screen "Balast Water Treatment Plant" 1280x800, template "Template"
   on GenerateScreen: "User_Change"(); "TitleUpdater"()
   Button "HmiScreenItemData_1" at 1,1 size 150x40; TextOn 'Back'; TextOff 'Main Index'
      on Release: ActivateScreen("02 Main Index", 0)
   TextField "Text field_63" at 383,107 size 72x30; Text 'Pre Dwell Time'
   Circle "Circle_29" at 1047,85 size 20x20
      Appearance <- "2102_TIME_CALCS_DB_POST_DWELL_TMR_DN"
   Button "HmiScreenItemData_9" at 10,60 size 158x27; TextOn 'Back'; TextOff 'BWTS Control'
   Button "HmiScreenItemData_4" at 14,150 size 75x47; TextOn 'Back'; TextOff 'Stop'; Authorization "Operate"
      on Release: function_efd93a16("BWTS Stop Confirm", 300, 200, -1, -1, 1)
      ObjectEnable <- "82_To_HMI_CRNT_MODE_GCU"
   Circle "Circle_20" at 137,105 size 29x29
      Appearance <- "80_From_HMI_RUN_IGG(1)"
   Button "HmiScreenItemData_3" at 14,93 size 75x47; TextOn 'Back'; TextOff 'Start'; Authorization "Operate"
      on Release: function_efd93a16("BWTS Start Confirm", 300, 200, -1, -1, 1)
      ObjectEnable <- "82_To_HMI_CRNT_MODE_GCU"
   Button "HmiScreenItemData_2" at 1129,1 size 150x40; TextOn 'Back'; TextOff 'BWTS Setup'
      on Release: ActivateScreen("Balast Water Treatment Setup", 0)
   TextField "Text field_1" at 290,107 size 68x30; Text 'Tank Selected'
   TextField "Text field_2" at 841,107 size 61x30; Text 'BWTS Started'
   TextField "Text field_3" at 568,107 size 62x30; Text 'IGGS Started'
   TextField "Text field_4" at 659,107 size 60x30; Text 'GCU Started'
   TextField "Text field_5" at 748,107 size 61x30; Text 'PGC Started'
   TextField "Text field_6" at 908,107 size 102x30; Text 'Gas Transfer Started'
   Circle "Circle_10" at 956,89 size 14x14
      Appearance <- "2110_BTCS_CNTRL_DB_BTCS_STEP"
   TextField "Text field_7" at 995,107 size 125x30; Text 'Treatment Cycle Completed'
   TextField "Text field_21" at 306,401 size 54x20; Text 'Closed'
      Visibility <- "20_TANKS_IP_DATA_RIO_06_FIRST_TANK_GTT_ISOL_VALVE_CLSD"
   TextField "Text field_22" at 306,401 size 54x20; Text 'Opened'
      Visibility <- "20_TANKS_IP_DATA_RIO_06_FIRST_TANK_GTT_ISOL_VALVE_OPEN"
   GraphicView "Graphic view_10" at 283,396 size 22x31; Picture "Graphic_162"
   TextField "Text field_25" at 306,482 size 54x20; Text 'Closed'
      Visibility <- "20_TANKS_IP_DATA_RIO_06_SECOND_TANK_GTT_ISOL_VALVE_CLSD"
   TextField "Text field_26" at 306,482 size 54x20; Text 'Opened'
      Visibility <- "20_TANKS_IP_DATA_RIO_06_SECOND_TANK_GTT_ISOL_VALVE_OPEN"
   IOField "I/O field_2" at 309,560 size 72x20; FormatPattern 999; Unit Nm³/hr
      ProcessValue <- "20_TANKS_IP_DATA_RIO_06_SECOND_TANK_USD_FLOW"
   IOField "I/O field_4" at 309,599 size 72x20; FormatPattern 999; Unit Nm³/hr
      ProcessValue <- "20_TANKS_IP_DATA_RIO_06_SECOND_TANK_MBG_FLOW"
   TextField "Text field_27" at 263,602 size 29x14; Text 'MBG'
   TextField "Text field_28" at 285,545 size 33x15; Text 'USD'
   TextField "Text field_23" at 261,291 size 34x14; Text 'MBG'
   TextField "Text field_24" at 284,349 size 28x14; Text 'USD'
   Group "Group" at 1064,419 size 35x38; Picture "Graphic_72"
   TextField "Text field_19" at 1057,414 size 54x20; Text 'Closed'
      Visibility <- "20_TANKS_IP_DATA_RIO_01_FIRST_TANK_GTT_ISOL_VALVE_CLSD"
   TextField "Text field_20" at 1057,414 size 54x20; Text 'Opened'
      Visibility <- "20_TANKS_IP_DATA_RIO_01_FIRST_TANK_GTT_ISOL_VALVE_OPEN"
   Group "Group_1" at 120,420 size 35x38; Picture "Graphic_72"
   TextField "Text field_72" at 112,415 size 54x20; Text 'Closed'
      Visibility <- "20_TANKS_IP_DATA_RIO_07_FIRST_TANK_GTT_ISOL_VALVE_CLSD"
   TextField "Text field_73" at 112,415 size 54x20; Text 'Opened'
      Visibility <- "20_TANKS_IP_DATA_RIO_07_FIRST_TANK_GTT_ISOL_VALVE_OPEN"
   TextField "Text field_8" at 438,401 size 54x20; Text 'Closed'
      Visibility <- "20_TANKS_IP_DATA_RIO_05_FIRST_TANK_GTT_ISOL_VALVE_CLSD"
   TextField "Text field_9" at 438,401 size 54x20; Text 'Opened'
      Visibility <- "20_TANKS_IP_DATA_RIO_05_FIRST_TANK_GTT_ISOL_VALVE_OPEN"
   GraphicView "Graphic view_1" at 415,396 size 22x31; Picture "Graphic_162"
   TextField "Text field_10" at 438,482 size 54x20; Text 'Closed'
      Visibility <- "20_TANKS_IP_DATA_RIO_05_SECOND_TANK_GTT_ISOL_VALVE_CLSD"
   TextField "Text field_11" at 438,482 size 54x20; Text 'Opened'
      Visibility <- "20_TANKS_IP_DATA_RIO_05_SECOND_TANK_GTT_ISOL_VALVE_OPEN"
   GraphicView "Graphic view_3" at 415,476 size 22x31; Picture "Graphic_162"
   IOField "I/O field_5" at 441,560 size 72x20; FormatPattern 999; Unit Nm³/hr
      ProcessValue <- "20_TANKS_IP_DATA_RIO_05_SECOND_TANK_USD_FLOW"
   IOField "I/O field_6" at 441,599 size 72x20; FormatPattern 999; Unit Nm³/hr
      ProcessValue <- "20_TANKS_IP_DATA_RIO_05_SECOND_TANK_MBG_FLOW"
   TextField "Text field_12" at 395,602 size 29x14; Text 'MBG'
   TextField "Text field_13" at 417,545 size 33x15; Text 'USD'
   IOField "I/O field_7" at 441,289 size 72x20; FormatPattern 999; Unit Nm³/hr
      ProcessValue <- "20_TANKS_IP_DATA_RIO_05_FIRST_TANK_MBG_FLOW"
   IOField "I/O field_8" at 441,330 size 72x20; FormatPattern 999; Unit Nm³/hr
      ProcessValue <- "20_TANKS_IP_DATA_RIO_05_FIRST_TANK_USD_FLOW"
   TextField "Text field_14" at 393,291 size 34x14; Text 'MBG'
   TextField "Text field_15" at 416,349 size 28x14; Text 'USD'
   TextField "Text field_16" at 570,402 size 54x20; Text 'Closed'
      Visibility <- "20_TANKS_IP_DATA_RIO_04_FIRST_TANK_GTT_ISOL_VALVE_CLSD"
   TextField "Text field_17" at 570,402 size 54x20; Text 'Opened'
      Visibility <- "20_TANKS_IP_DATA_RIO_04_FIRST_TANK_GTT_ISOL_VALVE_OPEN"
   GraphicView "Graphic view_15" at 547,396 size 22x31; Picture "Graphic_162"
   TextField "Text field_18" at 570,482 size 54x20; Text 'Closed'
      Visibility <- "20_TANKS_IP_DATA_RIO_04_SECOND_TANK_GTT_ISOL_VALVE_CLSD"
   TextField "Text field_29" at 570,482 size 54x20; Text 'Opened'
      Visibility <- "20_TANKS_IP_DATA_RIO_04_SECOND_TANK_GTT_ISOL_VALVE_OPEN"
   GraphicView "Graphic view_16" at 547,476 size 22x31; Picture "Graphic_162"
   IOField "I/O field_9" at 573,560 size 72x20; FormatPattern 999; Unit Nm³/hr
      ProcessValue <- "20_TANKS_IP_DATA_RIO_04_SECOND_TANK_USD_FLOW"
   IOField "I/O field_10" at 573,599 size 72x20; FormatPattern 999; Unit Nm³/hr
      ProcessValue <- "20_TANKS_IP_DATA_RIO_04_SECOND_TANK_MBG_FLOW"
   TextField "Text field_30" at 527,602 size 29x14; Text 'MBG'
   TextField "Text field_31" at 549,545 size 33x15; Text 'USD'
   IOField "I/O field_11" at 573,289 size 72x20; FormatPattern 999; Unit Nm³/hr
      ProcessValue <- "20_TANKS_IP_DATA_RIO_04_FIRST_TANK_MBG_FLOW"
   IOField "I/O field_12" at 573,330 size 72x20; FormatPattern 999; Unit Nm³/hr
      ProcessValue <- "20_TANKS_IP_DATA_RIO_04_FIRST_TANK_USD_FLOW"
   TextField "Text field_32" at 525,291 size 34x14; Text 'MBG'
   TextField "Text field_33" at 548,349 size 28x14; Text 'USD'
   TextField "Text field_34" at 702,401 size 54x20; Text 'Closed'
      Visibility <- "20_TANKS_IP_DATA_RIO_03_FIRST_TANK_GTT_ISOL_VALVE_CLSD"
   TextField "Text field_35" at 702,401 size 54x20; Text 'Opened'
      Visibility <- "20_TANKS_IP_DATA_RIO_03_FIRST_TANK_GTT_ISOL_VALVE_OPEN"
   GraphicView "Graphic view_21" at 679,396 size 22x31; Picture "Graphic_162"
   TextField "Text field_36" at 702,482 size 54x20; Text 'Closed'
      Visibility <- "20_TANKS_IP_DATA_RIO_03_SECOND_TANK_GTT_ISOL_VALVE_CLSD"
   TextField "Text field_37" at 702,482 size 54x20; Text 'Opened'
      Visibility <- "20_TANKS_IP_DATA_RIO_03_SECOND_TANK_GTT_ISOL_VALVE_OPEN"
   GraphicView "Graphic view_22" at 679,476 size 22x31; Picture "Graphic_162"
   IOField "I/O field_13" at 705,560 size 72x20; FormatPattern 999; Unit Nm³/hr
      ProcessValue <- "20_TANKS_IP_DATA_RIO_03_SECOND_TANK_USD_FLOW"
   IOField "I/O field_14" at 705,599 size 72x20; FormatPattern 999; Unit Nm³/hr
      ProcessValue <- "20_TANKS_IP_DATA_RIO_03_SECOND_TANK_MBG_FLOW"
   TextField "Text field_38" at 659,602 size 29x14; Text 'MBG'
   TextField "Text field_39" at 681,545 size 33x15; Text 'USD'
   IOField "I/O field_15" at 705,289 size 72x20; FormatPattern 999; Unit Nm³/hr
      ProcessValue <- "20_TANKS_IP_DATA_RIO_03_FIRST_TANK_MBG_FLOW"
   IOField "I/O field_16" at 705,330 size 72x20; FormatPattern 999; Unit Nm³/hr
      ProcessValue <- "20_TANKS_IP_DATA_RIO_03_FIRST_TANK_USD_FLOW"
   TextField "Text field_40" at 657,291 size 34x14; Text 'MBG'
   TextField "Text field_41" at 680,349 size 28x14; Text 'USD'
   TextField "Text field_42" at 834,401 size 54x20; Text 'Closed'
      Visibility <- "20_TANKS_IP_DATA_RIO_02_FIRST_TANK_GTT_ISOL_VALVE_CLSD"
   TextField "Text field_43" at 834,401 size 54x20; Text 'Opened'
      Visibility <- "20_TANKS_IP_DATA_RIO_02_FIRST_TANK_GTT_ISOL_VALVE_OPEN"
   GraphicView "Graphic view_27" at 811,396 size 22x31; Picture "Graphic_162"
   TextField "Text field_44" at 834,482 size 54x20; Text 'Closed'
      Visibility <- "20_TANKS_IP_DATA_RIO_02_SECOND_TANK_GTT_ISOL_VALVE_CLSD"
   TextField "Text field_45" at 834,482 size 54x20; Text 'Opened'
      Visibility <- "20_TANKS_IP_DATA_RIO_02_SECOND_TANK_GTT_ISOL_VALVE_OPEN"
   GraphicView "Graphic view_28" at 811,476 size 22x31; Picture "Graphic_162"
   IOField "I/O field_17" at 837,560 size 72x20; FormatPattern 999; Unit Nm³/hr
      ProcessValue <- "20_TANKS_IP_DATA_RIO_02_SECOND_TANK_USD_FLOW"
   IOField "I/O field_18" at 837,599 size 72x20; FormatPattern 999; Unit Nm³/hr
      ProcessValue <- "20_TANKS_IP_DATA_RIO_02_SECOND_TANK_MBG_FLOW"
   TextField "Text field_46" at 791,602 size 29x14; Text 'MBG'
   TextField "Text field_47" at 813,545 size 33x15; Text 'USD'
   IOField "I/O field_19" at 837,289 size 72x20; FormatPattern 999; Unit Nm³/hr
      ProcessValue <- "20_TANKS_IP_DATA_RIO_02_FIRST_TANK_MBG_FLOW"
   IOField "I/O field_20" at 837,330 size 72x20; FormatPattern 999; Unit Nm³/hr
      ProcessValue <- "20_TANKS_IP_DATA_RIO_02_FIRST_TANK_USD_FLOW"
   TextField "Text field_48" at 789,291 size 34x14; Text 'MBG'
   TextField "Text field_49" at 812,349 size 28x14; Text 'USD'
   TextField "Text field_50" at 966,401 size 54x20; Text 'Closed'
      Visibility <- "20_TANKS_IP_DATA_RIO_01_SECOND_TANK_GTT_ISOL_VALVE_CLSD"
   TextField "Text field_51" at 966,401 size 54x20; Text 'Opened'
      Visibility <- "20_TANKS_IP_DATA_RIO_01_SECOND_TANK_GTT_ISOL_VALVE_OPEN"
   GraphicView "Graphic view_33" at 943,396 size 22x31; Picture "Graphic_162"
   TextField "Text field_52" at 966,482 size 54x20; Text 'Closed'
      Visibility <- "20_TANKS_IP_DATA_RIO_01_THIRD_TANK_GTT_ISOL_VALVE_CLSD"
   TextField "Text field_53" at 966,482 size 54x20; Text 'Opened'
      Visibility <- "20_TANKS_IP_DATA_RIO_01_THIRD_TANK_GTT_ISOL_VALVE_OPEN"
   GraphicView "Graphic view_34" at 943,476 size 22x31; Picture "Graphic_162"
   IOField "I/O field_21" at 969,560 size 72x20; FormatPattern 999; Unit Nm³/hr
      ProcessValue <- "20_TANKS_IP_DATA_RIO_01_THIRD_TANK_USD_FLOW"
   IOField "I/O field_22" at 969,599 size 72x20; FormatPattern 999; Unit Nm³/hr
      ProcessValue <- "20_TANKS_IP_DATA_RIO_01_THIRD_TANK_MBG_FLOW"
   TextField "Text field_54" at 923,602 size 29x14; Text 'MBG'
   TextField "Text field_55" at 945,545 size 33x15; Text 'USD'
   IOField "I/O field_23" at 969,289 size 72x20; FormatPattern 999; Unit Nm³/hr
      ProcessValue <- "20_TANKS_IP_DATA_RIO_01_SECOND_TANK_MBG_FLOW"
   IOField "I/O field_24" at 969,330 size 72x20; FormatPattern 999; Unit Nm³/hr
      ProcessValue <- "20_TANKS_IP_DATA_RIO_01_SECOND_TANK_USD_FLOW"
   TextField "Text field_56" at 921,291 size 34x14; Text 'MBG'
   TextField "Text field_57" at 944,349 size 28x14; Text 'USD'
   GraphicView "Graphic view_17" at 575,446 size 485x12; Picture "Graphic_151"
   Button "Button_13" at 252,437 size 37x30; TextOff 'DB&B'
   TextField "Text field_58" at 188,226 size 50x40; Text 'Safe Area'
   TextField "Text field_59" at 417,454 size 137x22; Text 'Hazardous Area'
   IOField "I/O field_25" at 100,385 size 72x20; FormatPattern 999; Unit Nm³/hr
      ProcessValue <- "20_TANKS_IP_DATA_RIO_07_FIRST_TANK_MBG_FLOW"
   IOField "I/O field_26" at 100,491 size 72x20; FormatPattern 999; Unit Nm³/hr
      ProcessValue <- "20_TANKS_IP_DATA_RIO_07_FIRST_TANK_USD_FLOW"
   TextField "Text field_66" at 107,527 size 34x14; Text 'USD'
   TextField "Text field_67" at 107,356 size 34x14; Text 'MBG'
   IOField "I/O field_27" at 1073,381 size 72x20; FormatPattern 999; Unit Nm³/hr
      ProcessValue <- "20_TANKS_IP_DATA_RIO_01_FIRST_TANK_MBG_FLOW"
   IOField "I/O field_28" at 1080,491 size 72x20; FormatPattern 999; Unit Nm³/hr
      ProcessValue <- "20_TANKS_IP_DATA_RIO_01_FIRST_TANK_USD_FLOW"
   TextField "Text field_68" at 1111,527 size 34x14; Text 'USD'
   TextField "Text field_69" at 1111,350 size 34x14; Text 'MBG'
   Button "Button_20" at 724,152 size 115x34; TextOff 'Re-Oxygenation'
      Appearance <- "2110_BTCS_CNTRL_DB_BTCS_STEP"
   Button "Button_21" at 845,152 size 93x34; TextOff 'Post Dwell'
      Appearance <- "2110_BTCS_CNTRL_DB_BTCS_STATE"
   Circle "Circle_1" at 137,105 size 29x29
      Appearance <- "2110_BTCS_CNTRL_DB_BTCS_STATE"
   Circle "Circle_8" at 775,89 size 14x14
      Appearance <- "100_GCU_AUTO_SEQ_DB_CRNT_STEP"
   Circle "Circle_9" at 685,89 size 14x14
      Appearance <- "100_GCU_AUTO_SEQ_DB_CRNT_STEP"
   Circle "Circle_11" at 595,89 size 14x14
      Appearance <- "51_SLAVE_STATUS_RUNNING"
   Circle "Circle_12" at 866,89 size 14x14
      Appearance <- "2110_BTCS_CNTRL_DB_BTCS_STEP"
   Circle "Circle_13" at 324,89 size 14x14
      Appearance <- "HMI Indication Logic_DB_Tank Selected"
   Circle "Circle_14" at 414,89 size 14x14
      Appearance <- "2102_TIME_CALCS_DB_PRE_DWELL_TMR_DN"
   Button "Button_3" at 626,152 size 93x34; TextOff 'Dwell'
      Appearance <- "2110_BTCS_CNTRL_DB_BTCS_STATE"
   Button "Button_5" at 944,152 size 93x34; TextOff 'Complete'
      Appearance <- "HMI Indication Logic_DB_Sequence Finished"
   TextField "Text field_61" at 202,107 size 71x30; Text 'FA Mode Selected'
   Circle "Circle_2" at 230,89 size 14x14
      Appearance <- "HMI Indication Logic_DB_FA Mode Selected"
   TextField "Text field_60" at 190,519 size 46x25; Text 'GCU'
   GraphicIOField "Graphic I/O field_4" at 187,543 size 53x55; PictureList "GCU"
      ProcessValue <- "100_GCU_AUTO_SEQ_DB_RNG"
   TextField "Text field_65" at 190,398 size 46x25; Text 'PGC'
   TextField "Text field_74" at 186,279 size 54x25; Text 'IGGS'
   GraphicIOField "Graphic I/O field_1" at 185,303 size 57x53; PictureList "IGGS"
      ProcessValue <- "14_DQ_Data_24PF1"
   TextField "Text field_62" at 183,359 size 60x20; Text 'Disabled'
   TextField "Text field_77" at 183,359 size 60x20; Text 'Enabled'
      Visibility <- "51_SLAVE_STATUS_RUNNING"
   Button "Button_8" at 178,280 size 70x105; TextOff 'Text'
      on Release: ActivateScreen("Inert Gas Generator Plant", 0)
   TextField "Text field_75" at 183,480 size 60x20; Text 'Disabled'
   TextField "Text field_76" at 183,480 size 60x20; Text 'Enabled'
      Visibility <- "10_DI_DATA_E_400_RUN"
   TextField "Text field_70" at 183,599 size 60x20; Text 'Disabled'
   TextField "Text field_71" at 183,599 size 60x20; Text 'Enabled'
      Visibility <- "100_GCU_AUTO_SEQ_DB_RNG"
   Button "Button_4" at 178,521 size 70x105; TextOff 'Text'
      on Release: ActivateScreen("Inert Gas Conditioning Plant", 0)
   GraphicIOField "Graphic I/O field_2" at 770,45 size 250x30; PictureList "Process time Banner"
      ProcessValue <- "2110_BTCS_CNTRL_DB_BTCS_STATE"
      Visibility <- "2110_BTCS_CNTRL_DB_BTCS_STATE"
   Button "Button_14" at 303,152 size 93x34; TextOff 'Unselected'
      Visibility <- "HMI Indication Logic_DB_Tank Selected"
      Appearance <- "HMI Indication Logic_DB_Tank Selected"
   Button "Button_15" at 404,152 size 93x34; TextOff 'Selected'
      Appearance <- "HMI Indication Logic_DB_Tank Selected"
   Button "Button_16" at 506,152 size 115x34; TextOff 'De-Oxygenation'
      Appearance <- "2110_BTCS_CNTRL_DB_BTCS_STEP"
   TextField "Text field_78" at 115,457 size 55x26; Text 'CV-422 APT'
   GraphicView "Graphic view_76" at 185,421 size 57x55; Picture "Graphic_251"
   Button "Button_6" at 179,402 size 70x105; TextOff 'Text'
      on Release: ActivateScreen("PGC System", 0)
   TextField "Text field_79" at 297,421 size 71x15; Text 'CV-422-6P'
   TextField "Text field_80" at 429,421 size 71x15; Text 'CV-422-5P'
   TextField "Text field_81" at 561,421 size 71x15; Text 'CV-422-4P'
   TextField "Text field_82" at 693,421 size 71x15; Text 'CV-422-3P'
   TextField "Text field_83" at 825,421 size 71x15; Text 'CV-422-2P'
   TextField "Text field_84" at 957,421 size 71x15; Text 'CV-422-1P'
   TextField "Text field_85" at 1057,457 size 55x26; Text 'CV-422 FPT'
   TextField "Text field_86" at 297,503 size 70x15; Text 'CV-421-6S'
   TextField "Text field_87" at 429,503 size 70x15; Text 'CV-421-5S'
   TextField "Text field_88" at 561,503 size 70x15; Text 'CV-421-4S'
   TextField "Text field_89" at 693,503 size 70x15; Text 'CV-421-3S'
   TextField "Text field_90" at 825,503 size 70x15; Text 'CV-421-2S'
   TextField "Text field_91" at 957,503 size 70x15; Text 'CV-421-1S'
   TextField "Text field_93" at 436,351 size 76x15; Text 'FIT-418-5P'
   TextField "Text field_94" at 568,351 size 76x15; Text 'FIT-418-4P'
   TextField "Text field_95" at 700,351 size 76x15; Text 'FIT-418-3P'
   TextField "Text field_96" at 832,351 size 76x15; Text 'FIT-418-2P'
   TextField "Text field_97" at 964,351 size 76x15; Text 'FIT-418-1P'
   TextField "Text field_99" at 436,308 size 76x15; Text 'FIT-420-5P'
   TextField "Text field_100" at 568,308 size 76x15; Text 'FIT-420-4P'
   TextField "Text field_101" at 700,308 size 76x15; Text 'FIT-420-3P'
   TextField "Text field_102" at 832,308 size 76x15; Text 'FIT-420-2P'
   TextField "Text field_103" at 964,308 size 76x15; Text 'FIT-420-1P'
   TextField "Text field_104" at 90,369 size 85x15; Text 'FIT-420-APT'
   TextField "Text field_105" at 90,510 size 85x15; Text 'FIT-418-APT'
   TextField "Text field_106" at 1071,364 size 83x15; Text 'FIT-420-FPT'
   TextField "Text field_107" at 1071,510 size 83x15; Text 'FIT-418-FPT'
   TextField "Text field_108" at 304,620 size 75x15; Text 'FIT-419-6S'
   TextField "Text field_109" at 436,620 size 75x15; Text 'FIT-419-5S'
   TextField "Text field_110" at 568,620 size 75x15; Text 'FIT-419-4S'
   TextField "Text field_111" at 700,620 size 75x15; Text 'FIT-419-3S'
   TextField "Text field_112" at 832,620 size 75x15; Text 'FIT-419-2S'
   TextField "Text field_113" at 964,620 size 75x15; Text 'FIT-419-1S'
   TextField "Text field_114" at 304,579 size 75x15; Text 'FIT-417-6S'
   TextField "Text field_115" at 436,579 size 75x15; Text 'FIT-417-5S'
   TextField "Text field_116" at 568,579 size 75x15; Text 'FIT-417-4S'
   TextField "Text field_117" at 700,579 size 75x15; Text 'FIT-417-3S'
   TextField "Text field_118" at 832,579 size 75x15; Text 'FIT-417-2S'
   TextField "Text field_119" at 964,579 size 75x15; Text 'FIT-417-1S'
   Button "Button_63" at 1151,332 size 70x244; TextOff 'FPT'
      on Release: function_efd93a16("Tank FP Status", 168, 315, -1, 0, 1)
   Button "Button_24" at 1151,332 size 70x244; TextOff 'FPT'
      on Release: function_efd93a16("Tank FP Status", 168, 315, -1, 0, 1)
      Appearance <- "2110_BTCS_CNTRL_DB_BTCS_STATE"
      Visibility <- "504_Tank Grouping_DB2020_GROUP of TANK 1"
   Button "HmiScreenItemData_19" at 1185,676 size 72x27; TextOn 'Back'; TextOff 'Status'
      on Press: function_efd93a16("Treatment Status", 100, 471, -1, 3, 1)
   Group "Group_6" at 298,44 size 241x30
   Circle "Circle_26" at 504,89 size 14x14
      Appearance <- "2102_TIME_CALCS_DB_Time_To_Treatment"
   TextField "Text field_134" at 470,107 size 75x30; Text 'Wait for IGGS Start'
   GraphicView "Graphic view_26" at 1175,490 size 25x62; Picture "Graphic_183"
   GraphicView "Graphic view_29" at 1175,357 size 25x62; Picture "Graphic_183"
   Circle "Circle_24" at 1200,432 size 14x14
      Appearance <- "20_TANKS_IP_DATA_RIO_01_FIRST_TANK_BWT_LEVEL_HIHI"
   TextField "Text field_133" at 1171,432 size 35x14; Text 'LS425'
   Button "Button_64" at 921,206 size 124x70; TextOff 'Tank - 1P'
      on Release: function_efd93a16("Tank 1P Status", 168, 315, -1, 0, 1)
   Button "Button_22" at 921,206 size 124x70; TextOff 'Tank - 1P'
      on Release: function_efd93a16("Tank 1P Status", 168, 315, -1, 0, 1)
      Appearance <- "2110_BTCS_CNTRL_DB_BTCS_STATE"
      Visibility <- "504_Tank Grouping_DB2020_GROUP of TANK 2"
   Group "Group_3" at 925,210 size 117x62; Picture "Graphic_183"
   Button "Button_52" at 933,206 size 100x25; TextOff 'DISABLED'
      on Release: function_efd93a16("Tank 1P Status", 168, 315, -1, 0, 1)
      Visibility <- "504_Tank Grouping_DB2020_GROUP of TANK 2"
   Circle "Circle_16" at 999,253 size 14x14
      Appearance <- "20_TANKS_IP_DATA_RIO_01_SECOND_TANK_BWT_LEVEL_HIHI"
   TextField "Text field_120" at 955,253 size 51x14; Text 'LS425-1P'
   Button "Button_65" at 921,646 size 124x70; TextOff 'Tank - 1S'
      on Release: function_efd93a16("Tank 1S Status", 168, 315, -1, 0, 1)
   Button "Button_23" at 921,646 size 124x70; TextOff 'Tank - 1S'
      on Release: function_efd93a16("Tank 1S Status", 168, 315, -1, 0, 1)
      Appearance <- "2110_BTCS_CNTRL_DB_BTCS_STATE"
      Visibility <- "504_Tank Grouping_DB2020_GROUP of TANK 3"
   Group "Group_4" at 925,650 size 117x62; Picture "Graphic_183"
   Button "Button_54" at 933,691 size 100x25; TextOff 'DISABLED'
      on Release: function_efd93a16("Tank 1S Status", 168, 315, -1, 0, 1)
      Visibility <- "504_Tank Grouping_DB2020_GROUP of TANK 3"
   Circle "Circle_23" at 1000,653 size 14x14
      Appearance <- "20_TANKS_IP_DATA_RIO_01_THIRD_TANK_BWT_LEVEL_HIHI"
   TextField "Text field_126" at 955,654 size 51x14; Text 'LS422-1S'
   Button "Button_67" at 789,206 size 124x70; TextOff 'Tank - 2P'
      on Release: function_efd93a16("Tank 2P Status", 168, 315, -1, 0, 1)
   Button "Button_11" at 789,206 size 124x70; TextOff 'Tank - 2P'
      on Release: function_efd93a16("Tank 2P Status", 168, 315, -1, 0, 1)
      Appearance <- "2110_BTCS_CNTRL_DB_BTCS_STATE"
      Visibility <- "504_Tank Grouping_DB2020_GROUP of TANK 4"
   Group "Group_10" at 793,210 size 117x62; Picture "Graphic_183"
   Button "Button_32" at 801,206 size 100x25; TextOff 'DISABLED'
      on Release: function_efd93a16("Tank 2P Status", 168, 315, -1, 0, 1)
      Visibility <- "504_Tank Grouping_DB2020_GROUP of TANK 4"
   Circle "Circle_15" at 868,253 size 14x14
      Appearance <- "20_TANKS_IP_DATA_RIO_02_FIRST_TANK_BWT_LEVEL_HIHI"
   TextField "Text field_121" at 823,253 size 51x14; Text 'LS425-2P'
   Button "Button_69" at 789,646 size 124x70; TextOff 'Tank - 2S'
      on Release: function_efd93a16("Tank 2S Status", 168, 315, -1, 0, 1)
   Button "Button_7" at 789,646 size 124x70; TextOff 'Tank - 2S'
      on Release: function_efd93a16("Tank 2S Status", 168, 315, -1, 0, 1)
      Appearance <- "2110_BTCS_CNTRL_DB_BTCS_STATE"
      Visibility <- "504_Tank Grouping_DB2020_GROUP of TANK 5"
   Group "Group_13" at 793,650 size 117x62; Picture "Graphic_183"
   Button "Button_34" at 801,691 size 100x25; TextOff 'DISABLED'
      on Release: function_efd93a16("Tank 2S Status", 168, 315, -1, 0, 1)
      Visibility <- "504_Tank Grouping_DB2020_GROUP of TANK 5"
   Circle "Circle_22" at 868,653 size 14x14
      Appearance <- "20_TANKS_IP_DATA_RIO_02_SECOND_TANK_BWT_LEVEL_HIHI"
   TextField "Text field_127" at 823,654 size 51x14; Text 'LS422-2S'
   Button "Button_71" at 657,206 size 124x70; TextOff 'Tank - 3P'
      on Release: function_efd93a16("Tank 3P Status", 168, 315, -1, 0, 1)
   Button "Button_18" at 657,206 size 124x70; TextOff 'Tank - 3P'
      on Release: function_efd93a16("Tank 3P Status", 168, 315, -1, 0, 1)
      Appearance <- "2110_BTCS_CNTRL_DB_BTCS_STATE"
      Visibility <- "504_Tank Grouping_DB2020_GROUP of TANK 6"
   Group "Group_9" at 661,210 size 117x62; Picture "Graphic_183"
   Button "Button_36" at 669,206 size 100x25; TextOff 'DISABLED'
      on Release: function_efd93a16("Tank 3P Status", 168, 315, -1, 0, 1)
      Visibility <- "504_Tank Grouping_DB2020_GROUP of TANK 6"
   Circle "Circle_7" at 736,253 size 14x14
      Appearance <- "20_TANKS_IP_DATA_RIO_03_FIRST_TANK_BWT_LEVEL_HIHI"
   TextField "Text field_122" at 691,253 size 51x14; Text 'LS425-3P'
   Button "Button_73" at 657,646 size 124x70; TextOff 'Tank - 3S'
      on Release: function_efd93a16("Tank 3S Status", 168, 315, -1, 0, 1)
   Button "Button_9" at 657,646 size 124x70; TextOff 'Tank - 3S'
      on Release: function_efd93a16("Tank 3S Status", 168, 315, -1, 0, 1)
      Appearance <- "2110_BTCS_CNTRL_DB_BTCS_STATE"
      Visibility <- "504_Tank Grouping_DB2020_GROUP of TANK 7"
   Group "Group_12" at 661,650 size 117x62; Picture "Graphic_183"
   Button "Button_38" at 669,691 size 100x25; TextOff 'DISABLED'
      on Release: function_efd93a16("Tank 3S Status", 168, 315, -1, 0, 1)
      Visibility <- "504_Tank Grouping_DB2020_GROUP of TANK 7"
   Circle "Circle_21" at 736,653 size 14x14
      Appearance <- "20_TANKS_IP_DATA_RIO_03_SECOND_TANK_BWT_LEVEL_HIHI"
   TextField "Text field_128" at 691,654 size 51x14; Text 'LS422-3S'
   Button "Button_75" at 525,206 size 124x70; TextOff 'Tank - 4P'
      on Release: function_efd93a16("Tank 4P Status", 168, 315, -1, 2, 1)
   Button "Button_26" at 525,206 size 124x70; TextOff 'Tank - 4P'
      on Release: function_efd93a16("Tank 4P Status", 168, 315, -1, 2, 1)
      Appearance <- "2110_BTCS_CNTRL_DB_BTCS_STATE"
      Visibility <- "504_Tank Grouping_DB2020_GROUP of TANK 8"
   Group "Group_8" at 529,210 size 117x62; Picture "Graphic_183"
   Button "Button_40" at 537,206 size 100x25; TextOff 'DISABLED'
      on Release: function_efd93a16("Tank 4P Status", 168, 315, -1, 2, 1)
      Visibility <- "504_Tank Grouping_DB2020_GROUP of TANK 8"
   Circle "Circle_5" at 604,253 size 14x14
      Appearance <- "20_TANKS_IP_DATA_RIO_04_FIRST_TANK_BWT_LEVEL_HIHI"
   TextField "Text field_123" at 559,253 size 51x14; Text 'LS425-4P'
   Button "Button_80" at 393,646 size 124x70; TextOff 'Tank - 5S'
      on Release: function_efd93a16("Tank 5S Status", 168, 315, -1, 2, 1)
   Button "Button_25" at 393,646 size 124x70; TextOff 'Tank - 5S'
      on Release: function_efd93a16("Tank 5S Status", 168, 315, -1, 2, 1)
      Appearance <- "2110_BTCS_CNTRL_DB_BTCS_STATE"
      Visibility <- "504_Tank Grouping_DB2020_GROUP of TANK 11"
   GraphicView "Graphic view_13" at 489,650 size 25x62; Picture "Graphic_183"
   GraphicView "Graphic view_14" at 397,650 size 25x62; Picture "Graphic_183"
   Button "Button_46" at 405,691 size 100x25; TextOff 'DISABLED'
      on Release: function_efd93a16("Tank 5S Status", 168, 315, -1, 2, 1)
      Visibility <- "504_Tank Grouping_DB2020_GROUP of TANK 11"
   Circle "Circle_18" at 472,653 size 14x14
      Appearance <- "20_TANKS_IP_DATA_RIO_05_SECOND_TANK_BWT_LEVEL_HIHI"
   TextField "Text field_130" at 427,654 size 51x14; Text 'LS422-5S'
   Button "Button_81" at 525,646 size 124x70; TextOff 'Tank - 4S'
      on Release: function_efd93a16("Tank 4S Status", 168, 315, -1, 2, 1)
   Button "Button_19" at 525,646 size 124x70; TextOff 'Tank - 4S'
      on Release: function_efd93a16("Tank 4S Status", 168, 315, -1, 2, 1)
      Appearance <- "2110_BTCS_CNTRL_DB_BTCS_STATE"
      Visibility <- "504_Tank Grouping_DB2020_GROUP of TANK 9"
   Group "Group_11" at 529,650 size 117x62; Picture "Graphic_183"
   Button "Button_42" at 537,691 size 100x25; TextOff 'DISABLED'
      on Release: function_efd93a16("Tank 4S Status", 168, 315, -1, 2, 1)
      Visibility <- "504_Tank Grouping_DB2020_GROUP of TANK 9"
   Circle "Circle_19" at 604,653 size 14x14
      Appearance <- "20_TANKS_IP_DATA_RIO_04_SECOND_TANK_BWT_LEVEL_HIHI"
   TextField "Text field_129" at 559,654 size 51x14; Text 'LS422-4S'
   Button "Button_82" at 393,206 size 124x70; TextOff 'Tank - 5P'
      on Release: function_efd93a16("Tank 5P Status", 168, 315, -1, 2, 1)
   Button "Button_27" at 393,206 size 124x70; TextOff 'Tank - 5P'
      on Release: function_efd93a16("Tank 5P Status", 168, 315, -1, 2, 1)
      Appearance <- "2110_BTCS_CNTRL_DB_BTCS_STATE"
      Visibility <- "504_Tank Grouping_DB2020_GROUP of TANK 10"
   Group "Group_2" at 397,210 size 117x62; Picture "Graphic_183"
   Button "Button_44" at 405,206 size 100x25; TextOff 'DISABLED'
      on Release: function_efd93a16("Tank 5P Status", 168, 315, -1, 2, 1)
      Visibility <- "504_Tank Grouping_DB2020_GROUP of TANK 10"
   Circle "Circle_4" at 472,253 size 14x14
      Appearance <- "20_TANKS_IP_DATA_RIO_05_FIRST_TANK_BWT_LEVEL_HIHI"
   TextField "Text field_124" at 427,253 size 51x14; Text 'LS425-5P'
   Button "Button_83" at 261,206 size 124x70; TextOff 'Tank - 6P'
      on Release: function_efd93a16("Tank 6P Status", 168, 315, -1, 2, 1)
   Button "Button_28" at 261,206 size 124x70; TextOff 'Tank - 6P'
      on Release: function_efd93a16("Tank 6P Status", 168, 315, -1, 2, 1)
      Appearance <- "2110_BTCS_CNTRL_DB_BTCS_STATE"
      Visibility <- "504_Tank Grouping_DB2020_GROUP of TANK 12"
   GraphicView "Graphic view_4" at 357,210 size 25x62; Picture "Graphic_183"
   GraphicView "Graphic view_5" at 265,210 size 25x62; Picture "Graphic_183"
   Button "Button_48" at 273,206 size 100x25; TextOff 'DISABLED'
      on Release: function_efd93a16("Tank 6P Status", 168, 315, -1, 2, 1)
      Visibility <- "504_Tank Grouping_DB2020_GROUP of TANK 12"
   Circle "Circle_3" at 340,253 size 14x14
      Appearance <- "20_TANKS_IP_DATA_RIO_06_FIRST_TANK_BWT_LEVEL_HIHI"
   TextField "Text field_125" at 295,253 size 51x14; Text 'LS425-6P'
   Button "Button_85" at 261,646 size 124x70; TextOff 'Tank - 6S'
      on Release: function_efd93a16("Tank 6S Status", 168, 315, -1, 2, 1)
   Button "Button_29" at 261,646 size 124x70; TextOff 'Tank - 6S'
      on Release: function_efd93a16("Tank 6S Status", 168, 315, -1, 2, 1)
      Appearance <- "2110_BTCS_CNTRL_DB_BTCS_STATE"
      Visibility <- "504_Tank Grouping_DB2020_GROUP of TANK 13"
   GraphicView "Graphic view_7" at 357,650 size 25x62; Picture "Graphic_183"
   GraphicView "Graphic view_8" at 265,650 size 25x62; Picture "Graphic_183"
   Button "Button_50" at 273,691 size 100x25; TextOff 'DISABLED'
      on Release: function_efd93a16("Tank 6S Status", 168, 315, -1, 2, 1)
      Visibility <- "504_Tank Grouping_DB2020_GROUP of TANK 13"
   Circle "Circle_17" at 340,653 size 14x14
      Appearance <- "20_TANKS_IP_DATA_RIO_06_SECOND_TANK_BWT_LEVEL_HIHI"
   TextField "Text field_131" at 295,654 size 51x14; Text 'LS422-6S'
   Button "Button_87" at 51,369 size 45x172; TextOff 'APT'
      on Release: function_efd93a16("Tank AP Status", 168, 315, -1, 2, 1)
   Button "Button_1" at 51,369 size 45x172; TextOff 'APT'
      on Release: function_efd93a16("Tank AP Status", 168, 315, -1, 2, 1)
      Visibility <- "504_Tank Grouping_DB2020_GROUP of TANK 14"
      Appearance <- "2110_BTCS_CNTRL_DB_BTCS_STATE"
   GraphicView "Graphic view_30" at 62,383 size 21x46; Picture "Graphic_183"
   GraphicView "Graphic view_31" at 62,479 size 21x46; Picture "Graphic_183"
   Circle "Circle_25" at 79,432 size 14x14
      Appearance <- "20_TANKS_IP_DATA_RIO_07_FIRST_TANK_BWT_LEVEL_HIHI"
   TextField "Text field_132" at 50,432 size 35x14; Text 'LS425'
   IOField "I/O field_31" at 1053,45 size 225x30; FormatPattern ???????????????
      ProcessValue <- "Current User"
   Polyline "Polyline_1" at 261,205 size 123x70
      Visibility <- "504_Tank Grouping_DB2020_RUN TANK 12"
   Polyline "Polyline_2" at 392,205 size 123x70
      Visibility <- "504_Tank Grouping_DB2020_RUN TANK 10"
   Polyline "Polyline_3" at 525,205 size 123x70
      Visibility <- "504_Tank Grouping_DB2020_RUN TANK 8"
   Polyline "Polyline_4" at 656,205 size 123x70
      Visibility <- "504_Tank Grouping_DB2020_RUN TANK 6"
   Polyline "Polyline_5" at 789,205 size 123x70
      Visibility <- "504_Tank Grouping_DB2020_RUN TANK 4"
   Polyline "Polyline_6" at 921,205 size 123x70
      Visibility <- "504_Tank Grouping_DB2020_RUN TANK 2"
   Polyline "Polyline_7" at 921,646 size 123x70
      Visibility <- "504_Tank Grouping_DB2020_RUN TANK 3"
   Polyline "Polyline_8" at 789,646 size 123x70
      Visibility <- "504_Tank Grouping_DB2020_RUN TANK 5"
   Polyline "Polyline_9" at 658,646 size 123x70
      Visibility <- "504_Tank Grouping_DB2020_RUN TANK 7"
   Polyline "Polyline_10" at 525,646 size 123x70
      Visibility <- "504_Tank Grouping_DB2020_RUN TANK 9"
   Polyline "Polyline_11" at 393,646 size 123x70
      Visibility <- "504_Tank Grouping_DB2020_RUN TANK 11"
   GraphicView "Graphic view_12" at 283,476 size 22x31; Picture "Graphic_162"
   Polyline "Polyline_12" at 261,646 size 123x70
      Visibility <- "504_Tank Grouping_DB2020_RUN TANK 13"
   Polyline "Polyline_13" at 50,370 size 44x171
      Visibility <- "504_Tank Grouping_DB2020_RUN TANK 14"
   Button "Button_58" at 20,450 size 100x25; TextOff 'DISABLED'
      on Release: function_efd93a16("Tank AP Status", 168, 315, -1, 2, 1)
      Visibility <- "504_Tank Grouping_DB2020_GROUP of TANK 14"
   Polyline "Polyline_14" at 1152,332 size 68x242
      Visibility <- "504_Tank Grouping_DB2020_RUN TANK 1"
   Button "Button_56" at 1138,462 size 100x25; TextOff 'DISABLED'
      on Release: function_efd93a16("Tank FP Status", 168, 315, -1, 0, 1)
      Visibility <- "504_Tank Grouping_DB2020_GROUP of TANK 1"
   GraphicView "Graphic view_6" at 240,446 size 478x12; Picture "Graphic_151"
   Button "Button_2" at 252,437 size 37x30; TextOff 'DB&B'
      on Release: function_efd93a16("Double Block & Bleed Valve Monitoring", 250, 250, -1, -1, 1)
      Appearance <- "10_DI_DATA_CV407_OPN"
   Button "Button_84" at 258,203 size 126x73; TextOff 'Text'
      on Release: function_efd93a16("Tank 6P Status", 168, 315, -1, 0, 1)
      Appearance <- "504_Tank Grouping_DB2020_RUN TANK 12"
   Button "Button_76" at 524,204 size 126x73; TextOff 'Text'
      on Release: function_efd93a16("Tank 4P Status", 168, 315, -1, 0, 1)
      Appearance <- "504_Tank Grouping_DB2020_RUN TANK 8"
   Button "Button_72" at 655,204 size 126x73; TextOff 'Text'
      on Release: function_efd93a16("Tank 3P Status", 168, 315, -1, 0, 1)
      Appearance <- "504_Tank Grouping_DB2020_RUN TANK 6"
   Button "Button_68" at 787,204 size 126x73; TextOff 'Text'
      on Release: function_efd93a16("Tank 2P Status", 168, 315, -1, 0, 1)
      Appearance <- "504_Tank Grouping_DB2020_RUN TANK 4"
   Button "Button_62" at 920,203 size 126x73; TextOff 'Text'
      on Release: function_efd93a16("Tank 1P Status", 168, 315, -1, 0, 1)
      Appearance <- "504_Tank Grouping_DB2020_RUN TANK 2"
   Button "Button_61" at 1151,331 size 70x244; TextOff 'Text'
      on Release: function_efd93a16("Tank FP Status", 168, 315, -1, 0, 1)
      Appearance <- "504_Tank Grouping_DB2020_RUN TANK 1"
   Button "Button_88" at 49,369 size 47x174; TextOff 'Text'
      on Release: function_efd93a16("Tank AP Status", 168, 315, -1, 0, 1)
      Appearance <- "504_Tank Grouping_DB2020_RUN TANK 14"
   Button "Button_66" at 920,645 size 126x73; TextOff 'Text'
      on Release: function_efd93a16("Tank 1S Status", 168, 315, -1, 0, 1)
      Appearance <- "504_Tank Grouping_DB2020_RUN TANK 3"
   Button "Button_70" at 788,645 size 126x73; TextOff 'Text'
      on Release: function_efd93a16("Tank 2S Status", 168, 315, -1, 0, 1)
      Appearance <- "504_Tank Grouping_DB2020_RUN TANK 5"
   Button "Button_74" at 656,645 size 126x73; TextOff 'Text'
      on Release: function_efd93a16("Tank 3S Status", 168, 315, -1, 0, 1)
      Appearance <- "504_Tank Grouping_DB2020_RUN TANK 7"
   Button "Button_86" at 260,645 size 126x73; TextOff 'Text'
      on Release: function_efd93a16("Tank 6S Status", 168, 315, -1, 0, 1)
      Appearance <- "504_Tank Grouping_DB2020_RUN TANK 13"
   Button "Button_79" at 392,645 size 126x73; TextOff 'Text'
      on Release: function_efd93a16("Tank 5S Status", 168, 315, -1, 0, 1)
      Appearance <- "504_Tank Grouping_DB2020_RUN TANK 11"
   Button "Button_77" at 523,645 size 126x73; TextOff 'Text'
      on Release: function_efd93a16("Tank 4S Status", 168, 315, -1, 0, 1)
      Appearance <- "504_Tank Grouping_DB2020_RUN TANK 9"
   Button "HmiScreenItemData_8" at 920,732 size 355x40; TextOn 'Back'; TextOff 'Text'
   TextField "Screen title" at 906,728 size 373x50; Text 'Screen title'
   Button "HmiScreenItemData_6" at 1043,144 size 116x50; TextOn 'Back'; TextOff 'Tank Levels'
      on Release: ActivateScreen("Balast Water Treatment Plant Tank Levels", 0)
   GraphicView "Graphic view_107" at 302,354 size 64x55; Picture "Graphic_143"
      Visibility <- "2062_Warning_Data_Water Level Override 6P"
   IOField "I/O field_3" at 309,289 size 72x20; FormatPattern 999; Unit Nm³/hr
      ProcessValue <- "20_TANKS_IP_DATA_RIO_06_FIRST_TANK_MBG_FLOW"
   IOField "I/O field_1" at 309,330 size 72x20; FormatPattern 999; Unit Nm³/hr
      ProcessValue <- "20_TANKS_IP_DATA_RIO_06_FIRST_TANK_USD_FLOW"
   TextField "Text field_92" at 304,351 size 76x15; Text 'FIT-418-6P'
   TextField "Text field_98" at 304,308 size 76x15; Text 'FIT-420-6P'
   GraphicView "Graphic view_18" at 434,354 size 64x55; Picture "Graphic_143"
      Visibility <- "2062_Warning_Data_Water Level Override 5P"
   GraphicView "Graphic view_23" at 566,355 size 64x55; Picture "Graphic_143"
      Visibility <- "2062_Warning_Data_Water Level Override 4P"
   GraphicView "Graphic view_46" at 696,354 size 64x55; Picture "Graphic_143"
      Visibility <- "2062_Warning_Data_Water Level Override 3P"
   GraphicView "Graphic view_47" at 829,354 size 64x55; Picture "Graphic_143"
      Visibility <- "2062_Warning_Data_Water Level Override 2P"
   GraphicView "Graphic view_48" at 962,354 size 64x55; Picture "Graphic_143"
      Visibility <- "2062_Warning_Data_Water Level Override 1P"
   GraphicView "Graphic view_49" at 962,513 size 64x55; Picture "Graphic_143"
      Visibility <- "2062_Warning_Data_Water Level Override 1S"
   GraphicView "Graphic view_50" at 830,513 size 64x55; Picture "Graphic_143"
      Visibility <- "2062_Warning_Data_Water Level Override 2S"
   GraphicView "Graphic view_51" at 698,513 size 64x55; Picture "Graphic_143"
      Visibility <- "2062_Warning_Data_Water Level Override 3S"
   GraphicView "Graphic view_53" at 566,513 size 64x55; Picture "Graphic_143"
      Visibility <- "2062_Warning_Data_Water Level Override 4S"
   GraphicView "Graphic view_54" at 434,513 size 64x55; Picture "Graphic_143"
      Visibility <- "2062_Warning_Data_Water Level Override 5S"
   GraphicView "Graphic view_55" at 302,513 size 64x55; Picture "Graphic_143"
      Visibility <- "2062_Warning_Data_Water Level Override 6S"
   GraphicView "Graphic view_56" at 1153,283 size 64x55; Picture "Graphic_143"
      Visibility <- "2062_Warning_Data_Water Level Override FPT"
   GraphicView "Graphic view_57" at 41,321 size 64x55; Picture "Graphic_143"
      Visibility <- "2062_Warning_Data_Water Level Override APT"
   GraphicView "Graphic view_108" at 4,683 size 96x48; Picture "Left Arow"
   Button "HmiScreenItemData_14" at 3,660 size 106x93; TextOn 'Back'; TextOff 'Text'
      on Press: ActivateScreen("Inert Gas Conditioning Plant", 0)
   Button "Button_78" at 392,205 size 126x73; TextOff 'Text'
      on Release: function_efd93a16("Tank 5P Status", 168, 315, -1, 0, 1)
      Appearance <- "504_Tank Grouping_DB2020_RUN TANK 10"
   Group "Group_5" at 664,46 size 45x27; FormatPattern 999
   Group "Group_7" at 711,46 size 50x27; FormatPattern 999; Unit h
   Group "Group_14" at 605,46 size 57x27; FormatPattern 999; Unit h
   Button "HmiScreenItemData_5" at 180,144 size 116x50; TextOn 'Back'; TextOff 'Tank Status'
      on Release: function_efd93a16("Tank Status", 400, 250, -1, -1, 1)
   IOField "I/O field_36" at 1080,491 size 72x20; FormatPattern 999; Unit m³/hr
      ProcessValue <- "20_TANKS_IP_DATA_RIO_01_FIRST_TANK_USD FLOW  N"
      Visibility <- "Nm³/hr to m³/hr"
   IOField "I/O field_37" at 1073,381 size 72x20; FormatPattern 999; Unit m³/hr
      ProcessValue <- "20_TANKS_IP_DATA_RIO_01_FIRST_TANK_MBG_FLOW N"
      Visibility <- "Nm³/hr to m³/hr"
   IOField "I/O field_38" at 969,289 size 72x20; FormatPattern 999; Unit m³/hr
      ProcessValue <- "20_TANKS_IP_DATA_RIO_01_SECOND_TANK_MBG_FLOW N"
      Visibility <- "Nm³/hr to m³/hr"
   IOField "I/O field_39" at 969,330 size 72x20; FormatPattern 999; Unit m³/hr
      ProcessValue <- "20_TANKS_IP_DATA_RIO_01_SECOND_TANK_USD FLOW  N"
      Visibility <- "Nm³/hr to m³/hr"
   IOField "I/O field_40" at 969,560 size 72x20; FormatPattern 999; Unit m³/hr
      ProcessValue <- "20_TANKS_IP_DATA_RIO_01_THIRD_TANK_USD FLOW  N"
      Visibility <- "Nm³/hr to m³/hr"
   IOField "I/O field_41" at 969,599 size 72x20; FormatPattern 999; Unit m³/hr
      ProcessValue <- "20_TANKS_IP_DATA_RIO_01_THIRD_TANK_MBG_FLOW N"
      Visibility <- "Nm³/hr to m³/hr"
   IOField "I/O field_42" at 837,560 size 72x20; FormatPattern 999; Unit m³/hr
      ProcessValue <- "20_TANKS_IP_DATA_RIO_02_SECOND_TANK_USD FLOW  N"
      Visibility <- "Nm³/hr to m³/hr"
   IOField "I/O field_43" at 837,599 size 72x20; FormatPattern 999; Unit m³/hr
      ProcessValue <- "20_TANKS_IP_DATA_RIO_02_SECOND_TANK_MBG_FLOW N"
      Visibility <- "Nm³/hr to m³/hr"
   IOField "I/O field_44" at 837,289 size 72x20; FormatPattern 999; Unit m³/hr
      ProcessValue <- "20_TANKS_IP_DATA_RIO_02_FIRST_TANK_MBG_FLOW N"
      Visibility <- "Nm³/hr to m³/hr"
   IOField "I/O field_45" at 837,330 size 72x20; FormatPattern 999; Unit m³/hr
      ProcessValue <- "20_TANKS_IP_DATA_RIO_02_FIRST_TANK_USD FLOW  N"
      Visibility <- "Nm³/hr to m³/hr"
   IOField "I/O field_46" at 705,289 size 72x20; FormatPattern 999; Unit m³/hr
      ProcessValue <- "20_TANKS_IP_DATA_RIO_03_FIRST_TANK_MBG_FLOW N"
      Visibility <- "Nm³/hr to m³/hr"
   IOField "I/O field_47" at 705,330 size 72x20; FormatPattern 999; Unit m³/hr
      ProcessValue <- "20_TANKS_IP_DATA_RIO_03_FIRST_TANK_USD FLOW  N"
      Visibility <- "Nm³/hr to m³/hr"
   IOField "I/O field_48" at 705,560 size 72x20; FormatPattern 999; Unit m³/hr
      ProcessValue <- "20_TANKS_IP_DATA_RIO_03_SECOND_TANK_USD FLOW  N"
      Visibility <- "Nm³/hr to m³/hr"
   IOField "I/O field_49" at 705,599 size 72x20; FormatPattern 999; Unit m³/hr
      ProcessValue <- "20_TANKS_IP_DATA_RIO_03_SECOND_TANK_MBG_FLOW N"
      Visibility <- "Nm³/hr to m³/hr"
   IOField "I/O field_50" at 573,289 size 72x20; FormatPattern 999; Unit m³/hr
      ProcessValue <- "20_TANKS_IP_DATA_RIO_04_FIRST_TANK_MBG_FLOW N"
      Visibility <- "Nm³/hr to m³/hr"
   IOField "I/O field_51" at 573,330 size 72x20; FormatPattern 999; Unit m³/hr
      ProcessValue <- "20_TANKS_IP_DATA_RIO_04_FIRST_TANK_USD FLOW  N"
      Visibility <- "Nm³/hr to m³/hr"
   IOField "I/O field_52" at 573,560 size 72x20; FormatPattern 999; Unit m³/hr
      ProcessValue <- "20_TANKS_IP_DATA_RIO_04_SECOND_TANK_USD FLOW  N"
      Visibility <- "Nm³/hr to m³/hr"
   IOField "I/O field_53" at 573,599 size 72x20; FormatPattern 999; Unit m³/hr
      ProcessValue <- "20_TANKS_IP_DATA_RIO_04_SECOND_TANK_MBG_FLOW N"
      Visibility <- "Nm³/hr to m³/hr"
   IOField "I/O field_54" at 441,289 size 72x20; FormatPattern 999; Unit m³/hr
      ProcessValue <- "20_TANKS_IP_DATA_RIO_05_FIRST_TANK_MBG_FLOW N"
      Visibility <- "Nm³/hr to m³/hr"
   IOField "I/O field_55" at 441,330 size 72x20; FormatPattern 999; Unit m³/hr
      ProcessValue <- "20_TANKS_IP_DATA_RIO_05_FIRST_TANK_USD FLOW  N"
      Visibility <- "Nm³/hr to m³/hr"
   IOField "I/O field_56" at 441,560 size 72x20; FormatPattern 999; Unit m³/hr
      ProcessValue <- "20_TANKS_IP_DATA_RIO_05_SECOND_TANK_USD FLOW  N"
      Visibility <- "Nm³/hr to m³/hr"
   IOField "I/O field_57" at 441,599 size 72x20; FormatPattern 999; Unit m³/hr
      ProcessValue <- "20_TANKS_IP_DATA_RIO_05_SECOND_TANK_MBG_FLOW N"
      Visibility <- "Nm³/hr to m³/hr"
   IOField "I/O field_58" at 309,289 size 72x20; FormatPattern 999; Unit m³/hr
      ProcessValue <- "20_TANKS_IP_DATA_RIO_06_FIRST_TANK_MBG_FLOW N"
      Visibility <- "Nm³/hr to m³/hr"
   IOField "I/O field_59" at 309,330 size 72x20; FormatPattern 999; Unit m³/hr
      ProcessValue <- "20_TANKS_IP_DATA_RIO_06_FIRST_TANK_USD FLOW  N"
      Visibility <- "Nm³/hr to m³/hr"
   IOField "I/O field_60" at 309,560 size 72x20; FormatPattern 999; Unit m³/hr
      ProcessValue <- "20_TANKS_IP_DATA_RIO_06_SECOND_TANK_USD FLOW  N"
      Visibility <- "Nm³/hr to m³/hr"
   IOField "I/O field_61" at 309,599 size 72x20; FormatPattern 999; Unit m³/hr
      ProcessValue <- "20_TANKS_IP_DATA_RIO_06_SECOND_TANK_MBG_FLOW N"
      Visibility <- "Nm³/hr to m³/hr"
   IOField "I/O field_62" at 100,385 size 72x20; FormatPattern 999; Unit m³/hr
      ProcessValue <- "20_TANKS_IP_DATA_RIO_07_FIRST_TANK_MBG_FLOW N"
      Visibility <- "Nm³/hr to m³/hr"
   IOField "I/O field_63" at 100,491 size 72x20; FormatPattern 999; Unit m³/hr
      ProcessValue <- "20_TANKS_IP_DATA_RIO_07_FIRST_TANK_USD FLOW  N"
      Visibility <- "Nm³/hr to m³/hr"
   Button "HmiScreenItemData_7" at 1160,195 size 116x50; TextOn 'Back'; TextOff 'm³/hr to Nm³/hr Conversion'; TextList "m³/hr to Nm³/hr"
      ObjectEnable <- "user_group"
      Visibility <- "user_group"
      on Press: InvertBit("Nm³/hr to m³/hr")
      Appearance <- "Nm³/hr to m³/hr"
      ProcessValue <- "Nm³/hr to m³/hr"
   Button "Button_10" at 9,92 size 153x56; TextOff 'Text'
      on Release: function_efd93a16("Salinity - Acceptance", 168, 315, -1, 0, 1)
      Visibility <- "2068_Sys_Status_Data_SAL_VALID"
   Button "Button_12" at 9,92 size 153x57; TextOff 'Text'
      on Release: function_efd93a16("Tank Times", 300, 200, -1, 0, 1)
      Visibility <- "2068_Sys_Status_Data_Times Visibil"
   Button "HmiScreenItemData_10" at 1160,144 size 116x50; TextOn 'Back'; TextOff 'Tank Pressure'
      on Release: ActivateScreen("Balast Water Treatment Plant Tank Pressure", 0)
   GraphicView "Graphic view_52" at 1068,423 size 30x34; Picture "Graphic_72"
   GraphicView "Graphic view_2" at 124,424 size 30x34; Picture "Graphic_72"
   GraphicView "Graphic view_9" at 489,210 size 25x62; Picture "Graphic_183"
   GraphicView "Graphic view_11" at 397,210 size 25x62; Picture "Graphic_183"
   GraphicView "Graphic view_19" at 1017,210 size 25x62; Picture "Graphic_183"
   GraphicView "Graphic view_20" at 925,210 size 25x62; Picture "Graphic_183"
   GraphicView "Graphic view_24" at 1017,650 size 25x62; Picture "Graphic_183"
   GraphicView "Graphic view_25" at 925,650 size 25x62; Picture "Graphic_183"
   GraphicView "Graphic view_32" at 621,210 size 25x62; Picture "Graphic_183"
   GraphicView "Graphic view_35" at 529,210 size 25x62; Picture "Graphic_183"
   GraphicView "Graphic view_36" at 753,210 size 25x62; Picture "Graphic_183"
   GraphicView "Graphic view_37" at 661,210 size 25x62; Picture "Graphic_183"
   GraphicView "Graphic view_38" at 885,210 size 25x62; Picture "Graphic_183"
   GraphicView "Graphic view_39" at 793,210 size 25x62; Picture "Graphic_183"
   GraphicView "Graphic view_40" at 621,650 size 25x62; Picture "Graphic_183"
   GraphicView "Graphic view_41" at 529,650 size 25x62; Picture "Graphic_183"
   GraphicView "Graphic view_42" at 753,650 size 25x62; Picture "Graphic_183"
   GraphicView "Graphic view_43" at 661,650 size 25x62; Picture "Graphic_183"
   GraphicView "Graphic view_44" at 885,650 size 25x62; Picture "Graphic_183"
   GraphicView "Graphic view_45" at 793,650 size 25x62; Picture "Graphic_183"
   Button "Button_59" at 298,44 size 240x30; TextOn 'TB3 Enabled'; TextOff 'BWT System Shutting Down'
      Visibility <- "2110_BTCS_CNTRL_DB_BTCS_STATE"
   Button "Button_60" at 299,44 size 240x30; TextOn 'TB3 Enabled'; TextOff 'BWT System Enabled'
      Visibility <- "2110_BTCS_CNTRL_DB_BTCS_STATE"
   IOField "I/O field_29" at 664,46 size 45x27; FormatPattern 99; Unit h
      ProcessValue <- "Sequence Times_DB_Treatment Timer_Hours Left"
      Visibility <- "2110_BTCS_CNTRL_DB_BTCS_STATE"
   IOField "I/O field_30" at 664,46 size 45x27; FormatPattern 99; Unit h
      ProcessValue <- "Sequence Times_DB_Pre-Dwell Timer_Hours Left"
      Visibility <- "2110_BTCS_CNTRL_DB_BTCS_STATE"
   IOField "I/O field_32" at 711,46 size 50x27; FormatPattern 99; Unit m
      ProcessValue <- "Sequence Times_DB_Treatment Timer_Minutes Left"
      Visibility <- "2110_BTCS_CNTRL_DB_BTCS_STATE"
   IOField "I/O field_33" at 711,46 size 50x27; FormatPattern 99; Unit m
      ProcessValue <- "Sequence Times_DB_Pre-Dwell Timer_Minutes Left"
      Visibility <- "2110_BTCS_CNTRL_DB_BTCS_STATE"
   IOField "I/O field_34" at 605,46 size 57x27; FormatPattern 999; Unit d
      ProcessValue <- "Sequence Times_DB_Treatment Timer_Days Left"
      Visibility <- "2110_BTCS_CNTRL_DB_BTCS_STATE"
   IOField "I/O field_35" at 605,46 size 57x27; FormatPattern 999; Unit d
      ProcessValue <- "Sequence Times_DB_Pre-Dwell Timer_Days Left"
      Visibility <- "2110_BTCS_CNTRL_DB_BTCS_STATE"